(* Logix 5000 project; controller PLC_MCC1300_75F1 vendor 1 type 14 code 166 rev 32.11; software revision 32.04; part 7 of 83 *)

        [109].14   // Speed reference 3 M2CM10S
        [109].15   // Speed reference 4 M2CM10S
        [17].12   // VMCC TD SPARE
        [27].7   // Drive has a fault M2CM01
        [2].3   // VMCC M2 DC Output Power ON
        [113].0   // Drive ready M2CM11S
        [115].0   // Drive ready M2CM11N
        [117].0   // Drive ready M2CM12S
        [119].0   // Drive ready M2CM12N
        [123].11   // MB -->> M2 SPARE
        [31].7   // Drive has a fault M2CM3
        [102]   // RACK 14 INPUT UPDATES
        [104]   // Rack 15 Input Updates
        [1]   // RIO VMCC_TD_Inputs
        [17].13   // VMCC TD SPARE
        [49].11   // PANEL TD-CS4N SPARE
        [123].0   // MB -->> M2 SPARE
        [117].13   // Speed reference 2 M2CM12S
        [17].14   // VMCC TD SPARE
        [3].15   // VMCC M2 Drive fault Reset
        [53].13   // PANEL TD-CS5N SPARE
        [17].8   // VMCC TD Alarm Silence
        [2].10   // VMCC M2 E-STOP ACTIVE
        [2].5   // VMCC M2 E-STOP Power ON
        [32].12   // PANEL KD-CS1N SPARE
        [123].12   // MB -->> M2 SPARE
        [49].12   // PANEL TD-CS4N SPARE
        [106]   // Rack 15 Input Updates
        [108]   // Rack 15 Input Updates
        [17].15   // VMCC TD SPARE
        [49].13   // PANEL TD-CS4N SPARE
        [123].6   // MB -->> M2 SPARE
        [18].10   // VMCC TD SPARE
        [53].14   // PANEL TD-CS5N SPARE
        [53].15   // PANEL TD-CS5N SPARE
        [32].13   // PANEL KD-CS1N SPARE
        [32].14   // PANEL KD-CS1N SPARE
        [32].15   // PANEL KD-CS1N SPARE
        [33].10   // PANEL KD-CS1N SPARE
        [123].13   // MB -->> M2 SPARE
        [49].14   // PANEL TD-CS4N SPARE
        [110]   // Rack 15 Input Updates
        [112]   // Rack 16 Input Updates
        [18].11   // VMCC TD SPARE
        [49].15   // PANEL TD-CS4N SPARE
        [123].7   // MB -->> M2 SPARE
        [1].5   // Rockwell Run out Speed up signal M2CM7
        [117].14   // Speed reference 3 M2CM12S
        [123].8   // MB -->> M2 SPARE
        [117].15   // Speed reference 4 M2CM12S
        [117].2   // Command direction FW M2CM12S
        [117].3   // Actual direction FWD M2CM12S
        [33].0   // PANEL KD-CS1N Trim deck Move IN North Selector Sw.
        [36].2   // PANEL TD-CS1N Trim knocker 1 AUTO South Selector Sw.
        [117].6   // Drive has an alarm M2CM12S
        [117].7   // Drive has a fault M2CM12S
        [18].12   // VMCC TD SPARE
        [56].12   // PANEL TD-CS5S SPARE
        [56].13   // PANEL TD-CS5S SPARE
        [33].11   // PANEL KD-CS1N SPARE
        [33].12   // PANEL KD-CS1N SPARE
        [33].13   // PANEL KD-CS1N SPARE
        [33].14   // PANEL KD-CS1N SPARE
        [123].14   // MB -->> M2 SPARE
        [52].12   // PANEL TD-CS5N SPARE
        [114]   // Rack 16 Input Updates
        [116]   // Rack 16 Input Updates
        [18].13   // VMCC TD SPARE
        [52].13   // PANEL TD-CS5N SPARE
        [123].9   // MB -->> M2 SPARE
        [18].14   // VMCC TD SPARE
        [56].14   // PANEL TD-CS5S SPARE
        [57].10   // PANEL TD-CS5S SPARE
        [33].15   // PANEL KD-CS1N SPARE
        [37].11   // PANEL TD-CS1N SPARE
        [37].12   // PANEL TD-CS1N SPARE
        [37].13   // PANEL TD-CS1N SPARE
        [123].15   // MB -->> M2 SPARE
        [52].14   // PANEL TD-CS5N SPARE
        [118]   // Rack 16 Input Updates
        [120]   // Rack 17 Input Updates
        [18].15   // VMCC TD SPARE
        [52].15   // PANEL TD-CS5N SPARE
        [57].11   // PANEL TD-CS5S SPARE
        [57].12   // PANEL TD-CS5S SPARE
        [37].14   // PANEL TD-CS1N SPARE
        [37].15   // PANEL TD-CS1N SPARE
        [40].12   // PANEL TD-CS2N SPARE
        [40].13   // PANEL TD-CS2N SPARE
        [24].12   // I-SCAN BARS ON/OFF
        [53].10   // PANEL TD-CS5N SPARE
        [17].9   // VMCC TD Alarm Reset
        [29].1   // Drive running M2CM2
        [53].11   // PANEL TD-CS5N SPARE
        [1].6   // Rockwell Run out Speed up signal M2CM8
        [73].5   // BENCHBOARD Knurl Knocker Nth & Sth Auto mode
        [64].12   // Trim Deck PANEL TD-CS3S Crush all OFF Switch
        [73].7   // BENCHBOARD Knurl Knocker Master Auto mode
        [1].7   // Rockwell Run out Speed up signal M2CM9
        [37].7   // PANEL TD-CS1N Trim Conv 1 North Outer Limit Sw.
        [37].8   // PANEL TD-CS1N Trim Conv 1 North Inner Limit Sw.
        [33].8   // PANEL KD-CS1N Trim deck South Outer Limit Sw.
        [24].3   // RELIANCE CAPPING SYSTEM Trim Knocker #2 North Lower wheel
        [72].6   // BENCHBOARD Trim knocker #2 South Up Selector Sw.
        [72].8   // BENCHBOARD Trim knocker #3 North Up Selector Sw.
        [73].0   // BENCHBOARD Trim knocker #5 North Up Selector Sw.
        [24].15   // RELIANCE CAPPING SYSTEM Tracking window Lamp ON
        [33].4   // PANEL KD-CS1N Knurl knocker North Outer Limit Sw.
        [33].5   // PANEL KD-CS1N Knurl knocker North Inner Limit Sw.
        [33].9   // PANEL KD-CS1N Trim deck South Inner Limit Sw.
        [24].4   // RELIANCE CAPPING SYSTEM Trim Knocker #2 South Lower wheel
        [73].2   // BENCHBOARD Trim knocker #5 South Up Selector Sw.
        [37].10   // PANEL TD-CS1N Trim Conv 1 South Inner Limit Sw.
        [41].10   // PANEL TD-CS2N Trim Conv 2 North Outer Limit Sw.
        [41].11   // PANEL TD-CS2N Trim Conv 2 North Inner Limit Sw.
        [4].11   // VMCC M2 Speed zone 12 Drive Fault * 2CM12N
        [72].1   // BENCHBOARD Trim knocker #5 North Auto mode
        [72].3   // BENCHBOARD Trim knocker #5 South Auto mode
        [36].12   // PANEL TD-CS1N Float Glass Hold Down Wheels Auto Sel. Sw.
        [24].0   // RELIANCE CAPPING SYSTEM Knurl Knocker Nth & Sth Lower wheel
        [32].4   // PANEL KD-CS1N Knurl knocker Move UP South Selector Sw.
        [125].2   // ROCKWELL CAPPER Input to Disable manual y-cut bar 1
        [37].9   // PANEL TD-CS1N Trim Conv 1 South Outer Limit Sw.
        [36].1   // PANEL TD-CS1N Trim knocker 1 Move OUT South Selector Sw.
        [36].4   // PANEL TD-CS1N Trim knocker 1 Move UP South Selector Sw.
        [24].10   // RELIANCE CAPPING SYSTEM Trim Knocker #5 South Lower wheel
        [44].13   // Trim Deck PANEL TD-CS3N Crush all ON Switch
        [72].7   // BENCHBOARD Trim knocker #2 South Auto mode
        [45].6   // PANEL TD-CS3N Trim Conv 3 North Outer Limit Sw.
        [32].6   // PANEL KD-CS1N Knurl knocker Move IN North Selector Sw.
        [45].7   // PANEL TD-CS3N Trim Conv 3 North Inner Limit Sw.
        [72].9   // BENCHBOARD Trim knocker #3 North Auto mode
        [40].10   // PANEL TD-CS2N Trim knocker #2 Move UP North Selector Sw.
        [24].5   // RELIANCE CAPPING SYSTEM Trim Knocker #3 North Lower wheel
        [88]   // RACK 13 INPUT UPDATES
        [74]   // RACK 7 INPUT UPDATES
        [40].14   // PANEL TD-CS2N SPARE
        [24].6   // RELIANCE CAPPING SYSTEM Trim Knocker #3 South Lower wheel
        [90]   // RACK 13 INPUT UPDATES
        [103].14   // Speed reference 3 M2CM8N
        [119].10   // Local control 2 M2CM12N
        [109].2   // Command direction FW M2CM10S
        [115].12   // Speed reference 1 M2CM11N
        [36].8   // PANEL TD-CS1N Trim knocker 1 AUTO North Selector Sw.
        [36].14   // PANEL TD-CS1N Eclipse Hold Down Wheels Auto Sel. Sw.
        [36].3   // PANEL TD-CS1N Trim knocker 1 MANUAL South Selector Sw.
        [36].9   // PANEL TD-CS1N Trim knocker 1 MANUAL North Selector Sw.
        [69].5   // PANEL TD-CS2S Trim Conv 2 Move OUT North Selector Sw.
        [125].3   // ROCKWELL CAPPER Input to Disable auto y-cut bar 4
        [56].6   // PANEL TD-CS5S Trim knocker #5 Move IN North Selector Sw.
        [18].3   // VMCC TD SPARE
        [40].15   // PANEL TD-CS2N SPARE
        [41].14   // PANEL TD-CS2N SPARE
        [107].11   // Local control 3 M2CM9N
        [107].6   // Drive has an alarm M2CM9N
        [107].7   // Drive has a fault M2CM9N
        [105].9   // Local control 1 M2CM9S
        [41].15   // PANEL TD-CS2N SPARE
        [109].4   // Accelerating M2CM10S
        [2].8   // VMCC M2 Alarm Silence
        [31].1   // Drive running M2CM3
        [27].1   // Drive running M2CM01
        [18].5   // VMCC TD SPARE
        [44].14   // PANEL TD-CS3N SPARE
        [44].15   // PANEL TD-CS3N SPARE
        [109].10   // Local control 2 M2CM10S
        [109].11   // Local control 3 M2CM10S
        [109].7   // Drive has a fault M2CM10S
        [107].9   // Local control 1 M2CM9N
        [45].10   // PANEL TD-CS3N SPARE
        [109].5   // Decelerating M2CM10S
        [37].0   // PANEL TD-CS1N SPARE
        [37].1   // PANEL TD-CS1N SPARE
        [85].1   // Drive running M2CM4S
        [109].8   // Drive at speed M2CM10S
        [18].6   // VMCC TD SPARE
        [45].11   // PANEL TD-CS3N SPARE
        [45].12   // PANEL TD-CS3N SPARE
        [111].10   // Local control 2 M2CM10N
        [111].11   // Local control 3 M2CM10N
        [111].7   // Drive has a fault M2CM10N
        [111].8   // Drive at speed M2CM10N
        [45].13   // PANEL TD-CS3N SPARE
        [111].4   // Accelerating M2CM10N
        [37].4   // PANEL TD-CS1N SPARE
        [37].5   // PANEL TD-CS1N SPARE
        [87].1   // Drive running M2CM4N
        [18].7   // VMCC TD SPARE
        [45].14   // PANEL TD-CS3N SPARE
        [45].15   // PANEL TD-CS3N SPARE
        [113].10   // Local control 2 M2CM11S
        [113].11   // Local control 3 M2CM11S
        [113].7   // Drive has a fault M2CM11S
        [113].8   // Drive at speed M2CM11S
        [48].12   // PANEL TD-CS4N SPARE
        [111].5   // Decelerating M2CM10N
        [37].6   // PANEL TD-CS1N SPARE
        [4].12   // VMCC M2 Drive alarm
        [89].1   // Drive running M2CM5S
        [33].2   // PANEL KD-CS1N Trim deck Move IN South Selector Sw.
        [32].3   // PANEL KD-CS1N Knurl knocker MANUAL South Selector Sw.
        [73].14   // BENCHBOARD Input Power ON
        [57].13   // PANEL TD-CS5S SPARE
        [41].12   // PANEL TD-CS2N Trim Conv 2 South Outer Limit Sw.
        [36].11   // PANEL TD-CS1N Trim knocker 1 Move DOWN North Selector Sw.
        [3].9   // VMCC M2 Speed zone 10 Drive Fault 2CM10S
        [4].0   // VMCC M2 Speed zone 1 Drive Fault * 2CM01
        [4].1   // VMCC M2 Speed zone 2 Drive Fault * 2CM02
        [4].2   // VMCC M2 Speed zone 3 Drive Fault * 2CM03
        [73].3   // BENCHBOARD Knocker #5 South Auto mode
        [3].6   // VMCC M2 Speed zone 7 Drive Fault * 2CM07S
        [73].10   // Reliance BENCHBOARD Crush all OFF Switch
        [53].12   // PANEL TD-CS5N SPARE
        [113].4   // Accelerating M2CM11S
        [115].8   // Drive at speed M2CM11N
        [48].13   // PANEL TD-CS4N SPARE
        [73].15   // BENCHBOARD Output Power ON
        [117].8   // Drive at speed M2CM12S
        [36].13   // PANEL TD-CS1N Float Glass Hold Down Wheels Up Sel. Sw.
        [68].0   // PANEL TD-CS2S Trim knocker #2 Move IN South Selector Sw.
        [115].13   // Speed reference 2 M2CM11N
        [76].12   // PANEL KD-CS1S SPARE
        [40].5   // PANEL TD-CS2N Trim knocker #2 Move DOWN South Selector Sw.
        [44].10   // PANEL TD-CS3N Trim knocker #3 Move UP North Selector Sw.
        [44].5   // PANEL TD-CS3N Trim knocker #3 Move DOWN South Selector Sw.
        [24].7   // RELIANCE CAPPING SYSTEM Trim Knocker #4 North Lower wheel
        [103].2   // Command direction FW M2CM8N
        [125].4   // ROCKWELL CAPPER Input to Disable auto y-cut bar 3
        [103].15   // Speed reference 4 M2CM8N
        [2].0   // VMCC TD SPARE
        [81].0   // PANEL TD-CS1S SPARE
        [81].1   // PANEL TD-CS1S SPARE
        [57].14   // PANEL TD-CS5S SPARE
        [57].15   // PANEL TD-CS5S SPARE
        [60].12   // PANEL TD-CS4S SPARE
        [113].5   // Decelerating M2CM11S
        [81].4   // PANEL TD-CS1S SPARE
        [91].1   // Drive running M2CM5N
        [92]   // RACK 13 INPUT UPDATES
        [94]   // RACK 13 INPUT UPDATES
        [18].8   // VMCC TD SPARE
        [18].9   // VMCC TD SPARE
        [2].4   // VMCC M2 SPARE
        [81].5   // PANEL TD-CS1S SPARE
        [81].6   // PANEL TD-CS1S SPARE
        [60].13   // PANEL TD-CS4S SPARE
        [60].14   // PANEL TD-CS4S SPARE
        [60].15   // PANEL TD-CS4S SPARE
        [115].4   // Accelerating M2CM11N
        [93].1   // Drive running M2CM6S
        [96]   // RACK 14 INPUT UPDATES
        [98]   // RACK 14 INPUT UPDATES
        [2].13   // VMCC M2 SPARE
        [2].14   // VMCC M2 SPARE
        [3].0   // VMCC M2 SPARE
        [61].10   // PANEL TD-CS4S SPARE
        [61].11   // PANEL TD-CS4S SPARE
        [61].12   // PANEL TD-CS4S SPARE
        [115].5   // Decelerating M2CM11N
        [95].1   // Drive running M2CM6N
        [2].15   // VMCC M2 SPARE
        [3].12   // VMCC M2 SPARE
        [3].1   // VMCC M2 SPARE
        [61].13   // PANEL TD-CS4S SPARE
        [61].14   // PANEL TD-CS4S SPARE
        [61].15   // PANEL TD-CS4S SPARE
        [117].4   // Accelerating M2CM12S
        [97].1   // Drive running M2CM7S
        [3].13   // VMCC M2 SPARE
        [3].14   // VMCC M2 SPARE
        [3].2   // VMCC M2 SPARE
        [64].14   // PANEL TD-CS3S SPARE
        [64].15   // PANEL TD-CS3S SPARE
        [65].10   // PANEL TD-CS3S SPARE
        [117].5   // Decelerating M2CM12S
        [99].1   // Drive running M2CM7N
        [4].13   // VMCC M2 SPARE
        [4].14   // VMCC M2 SPARE
        [3].7   // VMCC M2 Speed zone 8 Drive Fault * 2CM08S
        [65].11   // PANEL TD-CS3S SPARE
        [65].12   // PANEL TD-CS3S SPARE
        [65].13   // PANEL TD-CS3S SPARE
        [119].4   // Accelerating M2CM12N
        [4].15   // VMCC M2 SPARE
        [64].13   // Trim Deck PANEL TD-CS3S Crush all ON Switch
        [41].13   // PANEL TD-CS2N Trim Conv 2 South Inner Limit Sw.
        [77].6   // PANEL KD-CS1S Trim deck North Outer Limit Sw.
        [45].8   // PANEL TD-CS3N Trim Conv 3 South Outer Limit Sw.
        [36].7   // PANEL TD-CS1N Trim knocker 1 Move OUT North Selector Sw.
        [69].10   // PANEL TD-CS2S Trim Conv 2 North Outer Limit Sw.
        [41].0   // PANEL TD-CS2N Trim Conv 1 Move IN North Selector Sw.
        [48].10   // PANEL TD-CS4N Trim knocker #4 Move UP North Selector Sw.
        [109].3   // Actual direction FWD M2CM10S
        [76].13   // PANEL KD-CS1S SPARE
        [109].6   // Drive has an alarm M2CM10S
        [40].0   // PANEL TD-CS2N Trim knocker #2 Move IN South Selector Sw.
        [32].9   // PANEL KD-CS1N Knurl knocker MANUAL North Selector Sw.
        [40].4   // PANEL TD-CS2N Trim knocker #2 Move UP South Selector Sw.
        [68].1   // PANEL TD-CS2S Trim knocker #2 Move OUT South Selector Sw.
        [52].1   // PANEL TD-CS5N Trim knocker #5 Move OUT South Selector Sw.
        [115].14   // Speed reference 3 M2CM11N
        [24].8   // RELIANCE CAPPING SYSTEM Trim Knocker #4 South Lower wheel
        [45].9   // PANEL TD-CS3N Trim Conv 3 South Inner Limit Sw.
        [69].7   // PANEL TD-CS2S Trim Conv 2 Move OUT South Selector Sw.
        [52].10   // PANEL TD-CS5N Trim knocker #5 Move UP North Selector Sw.
        [24].9   // RELIANCE CAPPING SYSTEM Trim Knocker #5 North Lower wheel
        [119].11   // Local control 3 M2CM12N
        [65].14   // PANEL TD-CS3S SPARE
        [76].14   // PANEL KD-CS1S SPARE
        [103].3   // Actual direction FWD M2CM8N
        [105].13   // Speed reference 2 M2CM9S
        [105].14   // Speed reference 3 M2CM9S
        [111].12   // Speed reference 1 M2CM10N
        [76].7   // PANEL KD-CS1S Knurl knocker Move OUT North Selector Sw.
        [80].0   // PANEL TD-CS1S Trim knocker 1 Move IN South Selector Sw.
        [119].12   // Speed reference 1 M2CM12N
        [105].15   // Speed reference 4 M2CM9S
        [111].13   // Speed reference 2 M2CM10N
        [119].13   // Speed reference 2 M2CM12N
        [40].11   // PANEL TD-CS2N Trim knocker #2 Move DOWN North Selector Sw.
        [56].7   // PANEL TD-CS5S Trim knocker #5 Move OUT North Selector Sw.
        [44].11   // PANEL TD-CS3N Trim knocker #3 Move DOWN North Selector Sw.
        [60].0   // PANEL TD-CS4S Trim knocker #4 Move IN South Selector Sw.
        [36].10   // PANEL TD-CS1N Trim knocker 1 Move UP North Selector Sw.
        [48].11   // PANEL TD-CS4N Trim knocker #4 Move DOWN North Selector Sw.
        [48].14   // PANEL TD-CS4N SPARE
        [105].12   // Speed reference 1 M2CM9S
        [69].11   // PANEL TD-CS2S Trim Conv 2 North Inner Limit Sw.
        [49].6   // PANEL TD-CS4N Trim Conv 4 North Outer Limit Sw.
        [48].15   // PANEL TD-CS4N SPARE
        [49].10   // PANEL TD-CS4N SPARE
        [60].1   // PANEL TD-CS4S Trim knocker #4 Move OUT South Selector Sw.
        [60].10   // PANEL TD-CS4S Trim knocker #4 Move UP North Selector Sw.
        [60].11   // PANEL TD-CS4S Trim knocker #4 Move DOWN North Selector Sw.
        [60].4   // PANEL TD-CS4S Trim knocker #4 Move UP South Selector Sw.
        [60].5   // PANEL TD-CS4S Trim knocker #4 Move DOWN South Selector Sw.
        [60].6   // PANEL TD-CS4S Trim knocker #4 Move IN North Selector Sw.
        [60].7   // PANEL TD-CS4S Trim knocker #4 Move OUT North Selector Sw.
        [76].15   // PANEL KD-CS1S SPARE
        [77].10   // PANEL KD-CS1S SPARE
        [77].11   // PANEL KD-CS1S SPARE
        [77].12   // PANEL KD-CS1S SPARE
        [77].13   // PANEL KD-CS1S SPARE
        [77].14   // PANEL KD-CS1S SPARE
        [77].15   // PANEL KD-CS1S SPARE
        [81].11   // PANEL TD-CS1S SPARE
        [81].12   // PANEL TD-CS1S SPARE
        [81].13   // PANEL TD-CS1S SPARE
        [81].14   // PANEL TD-CS1S SPARE
        [52].4   // PANEL TD-CS5N Trim knocker #5 Move UP South Selector Sw.
        [48].4   // PANEL TD-CS4N Trim knocker #4 Move UP South Selector Sw.
        [48].5   // PANEL TD-CS4N Trim knocker #4 Move DOWN South Selector Sw.
        [48].6   // PANEL TD-CS4N Trim knocker #4 Move IN North Selector Sw.
        [80].1   // PANEL TD-CS1S Trim knocker 1 Move OUT South Selector Sw.
        [41].2   // PANEL TD-CS2N Trim Conv 1 Move IN South Selector Sw.
        [40].2   // PANEL TD-CS2N Trim knocker #2 AUTO South Selector Sw.
        [40].8   // PANEL TD-CS2N Trim knocker #2 AUTO North Selector Sw.
        [119].14   // Speed reference 3 M2CM12N
        [69].12   // PANEL TD-CS2S Trim Conv 2 South Outer Limit Sw.
        [3].8   // VMCC M2 Speed zone 9 Drive Fault * 2CM09S
        [69].13   // PANEL TD-CS2S Trim Conv 2 South Inner Limit Sw.
        [4].3   // VMCC M2 Speed zone 4 Drive Fault * 2CM04N
        [77].4   // PANEL KD-CS1S Knurl knocker South Outer Limit Sw.
        [77].5   // PANEL KD-CS1S Knurl knocker South Inner Limit Sw.
        [4].4   // VMCC M2 Speed zone 5 Drive Fault * 2CM05N
        [80].15   // PANEL TD-CS1S Eclipse Hold Down Wheels Sel. Sw.
        [81].10   // PANEL TD-CS1S Trim Conv 1 South Inner Limit Sw.
        [4].5   // VMCC M2 Speed zone 6 Drive Fault * 2CM06N
        [4].6   // VMCC M2 Speed zone 7 Drive Fault * 2CM07N
        [4].7   // VMCC M2 Speed zone 8 Drive Fault * 2CM08N
        [4].8   // VMCC M2 Speed zone 9 Drive Fault * 2CM09N
        [4].9   // VMCC M2 Speed zone 10 Drive Fault * 2CM10
        [41].4   // PANEL TD-CS2N Trim Conv 2 Move IN North Selector Sw.
        [36].6   // PANEL TD-CS1N Trim knocker 1 Move IN North Selector Sw.
        [41].6   // PANEL TD-CS2N Trim Conv 2 Move IN South Selector Sw.
        [80].4   // PANEL TD-CS1S Trim knocker 1 Move UP South Selector Sw.
        [45].0   // PANEL TD-CS3N Trim Conv 3 Move IN North Selector Sw.
        [37].2   // PANEL TD-CS1N Trim knocker 1 North Outer Limit Sw.
        [40].3   // PANEL TD-CS2N Trim knocker #2 MANUAL South Selector Sw.
        [80].5   // PANEL TD-CS1S Trim knocker 1 Move DOWN South Selector Sw.
        [45].2   // PANEL TD-CS3N Trim Conv 3 Move IN South Selector Sw.
        [37].3   // PANEL TD-CS1N Trim knocker 1 North Inner Limit Sw.
        [49].0   // PANEL TD-CS4N Trim Conv 4 Move IN North Selector Sw.
        [72].10   // BENCHBOARD Trim knocker #3 South Up Selector Sw.
        [49].2   // PANEL TD-CS4N Trim Conv 4 Move IN South Selector Sw.
        [72].12   // BENCHBOARD Trim knocker #4 North Up Selector Sw.
        [53].0   // PANEL TD-CS5N Trim Conv 5 Move IN North Selector Sw.
        [72].14   // BENCHBOARD Trim knocker #4 South Up Selector Sw.
        [53].2   // PANEL TD-CS5N Trim Conv 5 Move IN South Selector Sw.
        [73].4   // BENCHBOARD Knurl Knocker Nth & Sth Up Selector Sw.
        [57].0   // PANEL TD-CS5S Trim Conv 5 Move IN North Selector Sw.
        [52].5   // PANEL TD-CS5N Trim knocker #5 Move DOWN South Selector Sw.
        [77].0   // PANEL KD-CS1S Trim deck Move IN North Selector Sw.
        [48].7   // PANEL TD-CS4N Trim knocker #4 Move OUT North Selector Sw.
        [40].9   // PANEL TD-CS2N Trim knocker #2 MANUAL North Selector Sw.
        [68].10   // PANEL TD-CS2S Trim knocker #2 Move UP North Selector Sw.
        [77].2   // PANEL KD-CS1S Trim deck Move IN South Selector Sw.
        [80].10   // PANEL TD-CS1S Trim knocker 1 Move UP North Selector Sw.
        [81].2   // PANEL TD-CS1S Trim knocker 1 South Outer Limit Sw.
        [57].2   // PANEL TD-CS5S Trim Conv 5 Move IN South Selector Sw.
        [52].11   // PANEL TD-CS5N Trim knocker #5 Move DOWN North Selector Sw.
        [56].1   // PANEL TD-CS5S Trim knocker #5 Move OUT South Selector Sw.
        [64].0   // PANEL TD-CS3S Trim knocker #3 Move IN South Selector Sw.
        [64].1   // PANEL TD-CS3S Trim knocker #3 Move OUT South Selector Sw.
        [64].10   // PANEL TD-CS3S Trim knocker #3 Move UP North Selector Sw.
        [64].11   // PANEL TD-CS3S Trim knocker #3 Move DOWN North Selector Sw.
        [36].5   // PANEL TD-CS1N Trim knocker 1 Move DOWN South Selector Sw.
        [119].15   // Speed reference 4 M2CM12N
        [40].1   // PANEL TD-CS2N Trim knocker #2 Move OUT South Selector Sw.
        [41].1   // PANEL TD-CS2N Trim Conv 1 Move OUT North Selector Sw.
        [41].3   // PANEL TD-CS2N Trim Conv 1 Move OUT South Selector Sw.
        [41].5   // PANEL TD-CS2N Trim Conv 2 Move OUT North Selector Sw.
        [41].7   // PANEL TD-CS2N Trim Conv 2 Move OUT South Selector Sw.
        [44].2   // PANEL TD-CS3N Trim knocker #3 AUTO South Selector Sw.
        [44].8   // PANEL TD-CS3N Trim knocker #3 AUTO North Selector Sw.
        [45].1   // PANEL TD-CS3N Trim Conv 3 Move OUT North Selector Sw.
        [52].6   // PANEL TD-CS5N Trim knocker #5 Move IN North Selector Sw.
        [64].4   // PANEL TD-CS3S Trim knocker #3 Move UP South Selector Sw.
        [64].5   // PANEL TD-CS3S Trim knocker #3 Move DOWN South Selector Sw.
        [40].7   // PANEL TD-CS2N Trim knocker #2 Move OUT North Selector Sw.
        [64].6   // PANEL TD-CS3S Trim knocker #3 Move IN North Selector Sw.
        [52].7   // PANEL TD-CS5N Trim knocker #5 Move OUT North Selector Sw.
        [44].3   // PANEL TD-CS3N Trim knocker #3 MANUAL South Selector Sw.
        [61].0   // PANEL TD-CS4S Trim Conv 4 Move IN North Selector Sw.
        [80].11   // PANEL TD-CS1S Trim knocker 1 Move DOWN North Selector Sw.
        [56].10   // PANEL TD-CS5S Trim knocker #5 Move UP North Selector Sw.
        [80].6   // PANEL TD-CS1S Trim knocker 1 Move IN North Selector Sw.
        [68].11   // PANEL TD-CS2S Trim knocker #2 Move DOWN North Selector Sw.
        [56].0   // PANEL TD-CS5S Trim knocker #5 Move IN South Selector Sw.
        [44].9   // PANEL TD-CS3N Trim knocker #3 MANUAL North Selector Sw.
        [81].15   // PANEL TD-CS1S SPARE
        [61].2   // PANEL TD-CS4S Trim Conv 4 Move IN South Selector Sw.
        [65].0   // PANEL TD-CS3S Trim Conv 3 Move IN North Selector Sw.
        [64].7   // PANEL TD-CS3S Trim knocker #3 Move OUT North Selector Sw.
        [56].11   // PANEL TD-CS5S Trim knocker #5 Move DOWN North Selector Sw.
        [80].12   // PANEL TD-CS1S Float Glass Hold Down Wheels Auto Sel. Sw.
        [45].3   // PANEL TD-CS3N Trim Conv 3 Move OUT South Selector Sw.
        [80].13   // PANEL TD-CS1S Float Glass Hold Down Wheels Up Sel. Sw.
        [68].4   // PANEL TD-CS2S Trim knocker #2 Move UP South Selector Sw.
        [80].7   // PANEL TD-CS1S Trim knocker 1 Move OUT North Selector Sw.
        [49].7   // PANEL TD-CS4N Trim Conv 4 North Inner Limit Sw.
        [49].8   // PANEL TD-CS4N Trim Conv 4 South Outer Limit Sw.
        [49].9   // PANEL TD-CS4N Trim Conv 4 South Inner Limit Sw.
        [53].6   // PANEL TD-CS5N Trim Conv 5 North Outer Limit Sw.
        [53].7   // PANEL TD-CS5N Trim Conv 5 North Inner Limit Sw.
        [57].6   // PANEL TD-CS5S Trim Conv 5 North Outer Limit Sw.
        [57].7   // PANEL TD-CS5S Trim Conv 5 North Inner Limit Sw.
        [57].8   // PANEL TD-CS5S Trim Conv 5 South Outer Limit Sw.
        [57].9   // PANEL TD-CS5S Trim Conv 5 South Inner Limit Sw.
        [61].6   // PANEL TD-CS4S Trim Conv 4 North Outer Limit Sw.
        [81].3   // PANEL TD-CS1S Trim knocker 1 South Inner Limit Sw.
        [119].2   // Command direction FW M2CM12N
        [85].7   // Drive has a fault M2CM4S
        [44].1   // PANEL TD-CS3N Trim knocker #3 Move OUT South Selector Sw.
        [61].7   // PANEL TD-CS4S Trim Conv 4 North Inner Limit Sw.
        [61].8   // PANEL TD-CS4S Trim Conv 4 South Outer Limit Sw.
        [48].3   // PANEL TD-CS4N Trim knocker #4 MANUAL South Selector Sw.
        [48].2   // PANEL TD-CS4N Trim knocker #4 AUTO South Selector Sw.
        [87].7   // Drive has a fault M2CM4N
        [61].9   // PANEL TD-CS4S Trim Conv 4 South Inner Limit Sw.
        [89].7   // Drive has a fault M2CM5S
        [68].5   // PANEL TD-CS2S Trim knocker #2 Move DOWN South Selector Sw.
        [48].8   // PANEL TD-CS4N Trim knocker #4 AUTO North Selector Sw.
        [65].6   // PANEL TD-CS3S Trim Conv 3 North Outer Limit Sw.
        [119].3   // Actual direction FWD M2CM12N
        [68].6   // PANEL TD-CS2S Trim knocker #2 Move IN North Selector Sw.
        [65].2   // PANEL TD-CS3S Trim Conv 3 Move IN South Selector Sw.
        [44].6   // PANEL TD-CS3N Trim knocker #3 Move IN North Selector Sw.
        [40].6   // PANEL TD-CS2N Trim knocker #2 Move IN North Selector Sw.
        [119].6   // Drive has an alarm M2CM12N
        [44].0   // PANEL TD-CS3N Trim knocker #3 Move IN South Selector Sw.
        [68].7   // PANEL TD-CS2S Trim knocker #2 Move OUT North Selector Sw.
        [69].0   // PANEL TD-CS2S Trim Conv 1 Move IN North Selector Sw.
        [44].7   // PANEL TD-CS3N Trim knocker #3 Move OUT North Selector Sw.
        [65].7   // PANEL TD-CS3S Trim Conv 3 North Inner Limit Sw.
        [65].8   // PANEL TD-CS3S Trim Conv 3 South Outer Limit Sw.
        [65].9   // PANEL TD-CS3S Trim Conv 3 South Inner Limit Sw.
        [73].6   // BENCHBOARD Knurl Knocker Master Up Selector Sw.
        [81].7   // PANEL TD-CS1S Trim Conv 1 North Outer Limit Sw.
        [81].8   // PANEL TD-CS1S Trim Conv 1 North Inner Limit Sw.
        [81].9   // PANEL TD-CS1S Trim Conv 1 South Outer Limit Sw.
        [48].0   // PANEL TD-CS4N Trim knocker #4 Move IN South Selector Sw.
        [77].7   // PANEL KD-CS1S Trim deck North Inner Limit Sw.
        [77].8   // PANEL KD-CS1S Trim deck South Outer Limit Sw.
        [77].9   // PANEL KD-CS1S Trim deck South Inner Limit Sw.
        [52].0   // PANEL TD-CS5N Trim knocker #5 Move IN South Selector Sw.
        [91].7   // Drive has a fault M2CM5N
        [93].7   // Drive has a fault M2CM6S
        [95].7   // Drive has a fault M2CM6N
        [97].7   // Drive has a fault M2CM7S
        [69].2   // PANEL TD-CS2S Trim Conv 1 Move IN South Selector Sw.
        [56].4   // PANEL TD-CS5S Trim knocker #5 Move UP South Selector Sw.
        [49].1   // PANEL TD-CS4N Trim Conv 4 Move OUT North Selector Sw.
        [125].5   // ROCKWELL CAPPER Input to Disable auto y-cut bar 2
        [125].6   // ROCKWELL CAPPER Input to Disable auto y-cut bar 1
        [32].2   // PANEL KD-CS1N Knurl knocker AUTO South Selector Sw.
        [32].8   // PANEL KD-CS1N Knurl knocker AUTO North Selector Sw.
        [33].1   // PANEL KD-CS1N Trim deck Move OUT North Selector Sw.
        [33].3   // PANEL KD-CS1N Trim deck Move OUT South Selector Sw.
        [41].8   // PANEL TD-CS2N Trim knocker #2 North Outer Limit Sw.
        [41].9   // PANEL TD-CS2N Trim knocker #2 North Inner Limit Sw.
        [45].4   // PANEL TD-CS3N Trim knocker #3 North Outer Limit Sw.
        [45].5   // PANEL TD-CS3N Trim knocker #3 North Inner Limit Sw.
        [49].4   // PANEL TD-CS4N Trim knocker #4 North Outer Limit Sw.
        [49].5   // PANEL TD-CS4N Trim knocker #4 North Inner Limit Sw.
        [53].8   // PANEL TD-CS5S Trim knocker #5 South Outer Limit Sw.
        [53].9   // PANEL TD-CS5S Trim knocker #5 South Inner Limit Sw.
        [61].4   // PANEL TD-CS4S Trim knocker #4 South Outer Limit Sw.
        [61].5   // PANEL TD-CS4S Trim knocker #4 South Inner Limit Sw.
        [65].4   // PANEL TD-CS3S Trim knocker #3 South Outer Limit Sw.
        [99].7   // Drive has a fault M2CM7N
        [119].7   // Drive has a fault M2CM12N
        [17].11   // VMCC TD Panel Overtemp Alarm
        [17].3   // VMCC TD DC Output Power ON
        [17].4   // VMCC TD DC Power Supply #1 ON
        [76].10   // PANEL KD-CS1S Knurl knocker Move UP North Selector Sw.
        [49].3   // PANEL TD-CS4N Trim Conv 4 Move OUT South Selector Sw.
        [76].0   // PANEL KD-CS1S Knurl knocker Move IN South Selector Sw.
        [76].3   // PANEL KD-CS1S Knurl knocker MANUAL South Selector Sw.
        [76].4   // PANEL KD-CS1S Knurl knocker Move UP South Selector Sw.
        [76].6   // PANEL KD-CS1S Knurl knocker Move IN North Selector Sw.
        [17].6   // VMCC TD DC Power Supply #2 ON
        [52].2   // PANEL TD-CS5N Trim knocker #5 AUTO South Selector Sw.
        [52].8   // PANEL TD-CS5N Trim knocker #5 AUTO North Selector Sw.
        [69].4   // PANEL TD-CS2S Trim Conv 2 Move IN North Selector Sw.
        [65].5   // PANEL TD-CS3S Trim knocker #3 South Inner Limit Sw.
        [69].8   // PANEL TD-CS2S Trim knocker #2 South Outer Limit Sw.
        [53].1   // PANEL TD-CS5N Trim Conv 5 Move OUT North Selector Sw.
        [53].3   // PANEL TD-CS5N Trim Conv 5 Move OUT South Selector Sw.
        [69].6   // PANEL TD-CS2S Trim Conv 2 Move IN South Selector Sw.
        [69].9   // PANEL TD-CS2S Trim knocker #2 South Inner Limit Sw.
        [76].2   // PANEL KD-CS1S Knurl knocker AUTO South Selector Sw.
        [56].2   // PANEL TD-CS5S Trim knocker #5 AUTO South Selector Sw.
        [56].8   // PANEL TD-CS5S Trim knocker #5 AUTO North Selector Sw.
        [80].2   // PANEL TD-CS1S Trim knocker 1 AUTO South Selector Sw.
        [76].8   // PANEL KD-CS1S Knurl knocker AUTO North Selector Sw.
        [77].1   // PANEL KD-CS1S Trim deck Move OUT North Selector Sw.
        [57].1   // PANEL TD-CS5S Trim Conv 5 Move OUT North Selector Sw.
        [57].3   // PANEL TD-CS5S Trim Conv 5 Move OUT South Selector Sw.
        [80].8   // PANEL TD-CS1S Trim knocker 1 AUTO North Selector Sw.
        [77].3   // PANEL KD-CS1S Trim deck Move OUT South Selector Sw.
        [48].9   // PANEL TD-CS4N Trim knocker #4 MANUAL North Selector Sw.
        [52].3   // PANEL TD-CS5N Trim knocker #5 MANUAL South Selector Sw.
        [76].9   // PANEL KD-CS1S Knurl knocker MANUAL North Selector Sw.
        [60].2   // PANEL TD-CS4S Trim knocker #4 AUTO South Selector Sw.
        [60].8   // PANEL TD-CS4S Trim knocker #4 AUTO North Selector Sw.
        [52].9   // PANEL TD-CS5N Trim knocker #5 MANUAL North Selector Sw.
        [56].3   // PANEL TD-CS5S Trim knocker #5 MANUAL South Selector Sw.
        [80].14   // PANEL TD-CS1S Eclipse Hold Down Wheels Auto Sel. Sw.
        [61].1   // PANEL TD-CS4S Trim Conv 4 Move OUT North Selector Sw.
        [61].3   // PANEL TD-CS4S Trim Conv 4 Move OUT South Selector Sw.
        [56].9   // PANEL TD-CS5S Trim knocker #5 MANUAL North Selector Sw.
        [60].3   // PANEL TD-CS4S Trim knocker #4 MANUAL South Selector Sw.
        [80].3   // PANEL TD-CS1S Trim knocker 1 MANUAL South Selector Sw.
        [64].2   // PANEL TD-CS3S Trim knocker #3 AUTO South Selector Sw.
        [64].8   // PANEL TD-CS3S Trim knocker #3 AUTO North Selector Sw.
        [60].9   // PANEL TD-CS4S Trim knocker #4 MANUAL North Selector Sw.
        [64].3   // PANEL TD-CS3S Trim knocker #3 MANUAL South Selector Sw.
        [80].9   // PANEL TD-CS1S Trim knocker 1 MANUAL North Selector Sw.
        [65].1   // PANEL TD-CS3S Trim Conv 3 Move OUT North Selector Sw.
        [65].3   // PANEL TD-CS3S Trim Conv 3 Move OUT South Selector Sw.
        [64].9   // PANEL TD-CS3S Trim knocker #3 MANUAL North Selector Sw.
        [68].3   // PANEL TD-CS2S Trim knocker #2 MANUAL South Selector Sw.
        [68].2   // PANEL TD-CS2S Trim knocker #2 AUTO South Selector Sw.
        [68].8   // PANEL TD-CS2S Trim knocker #2 AUTO North Selector Sw.
        [68].9   // PANEL TD-CS2S Trim knocker #2 MANUAL North Selector Sw.
        [76].1   // PANEL KD-CS1S Knurl knocker Move OUT South Selector Sw.
        [69].1   // PANEL TD-CS2S Trim Conv 1 Move OUT North Selector Sw.
        [69].3   // PANEL TD-CS2S Trim Conv 1 Move OUT South Selector Sw.
        [44].4   // PANEL TD-CS3N Trim knocker #3 Move UP South Selector Sw.
        [17].7   // VMCC TD DC Power Supply #3 ON
        [48].1   // PANEL TD-CS4N Trim knocker #4 Move OUT South Selector Sw.
   KD_N_MOVIN : ALIAS FOR N14[256].0;
   KD_N_MOVOUT : ALIAS FOR N14[257].0;
   KD_S_MOVIN : ALIAS FOR N14[256].1;
   KD_S_MOVOUT : ALIAS FOR N14[257].1;
   KK_N_MOVDN : ALIAS FOR N14[253].0;
   KK_N_MOVIN : ALIAS FOR N14[254].0;
   KK_N_MOVOUT : ALIAS FOR N14[255].0;
   KK_N_MOVUP : ALIAS FOR N14[252].0;
   KK_S_MOVDN : ALIAS FOR N14[253].1;
   KK_S_MOVIN : ALIAS FOR N14[254].1;
   KK_S_MOVOUT : ALIAS FOR N14[255].1;
   KK_S_MOVUP : ALIAS FOR N14[252].1;
   KNRL_K_NTH_ADJ : ALIAS FOR O[19].0;
   KNRL_K_STH_ADJ : ALIAS FOR O[19].1;
   KNRL_N_AUTO : ALIAS FOR N14[250].0;
   KNRL_N_MANL : ALIAS FOR N14[251].0;
   KNRL_S_AUTO : ALIAS FOR N14[250].1;
   KNRL_S_MANL : ALIAS FOR N14[251].1;
   KNRL_T_NTH_ADJ : ALIAS FOR O[22].0;
   KNRL_T_STH_ADJ : ALIAS FOR O[22].1;
   LEHR_SPEED : ALIAS FOR N20[1];
   LINE_SPEED : ALIAS FOR N20[3];
   M2_ALM_HORN_RLY : ALIAS FOR O[9].3;
   M2_ALM_RESET : ALIAS FOR I[2].9;
   M2_ALM_SILENCE : ALIAS FOR I[2].8;
   M2_AMBER_STKLTE : ALIAS FOR O[9].6;
   M2_BLUE_STKLTE : ALIAS FOR O[9].5;
   M2_CM07N_HZIMP : DINT := 1853;   // This compute statement was created to allow speed control on M2 CM07N; 28Mar2019,AAC.
   M2_CM07N_Lehr_Speed : DINT := 71;   // This compute statement was created to allow speed control for Lehr Speed on M2 CM07N; 28Mar2019,AAC.
   M2_CM07N_Slip_Comp : DINT := 1160;
   M2_CM07N_Trim_Speed : DINT := 243;   // This compute statement was created to allow Trim speed control on M2 CM07N; 28Mar2019,AAC.
   M2_DC_INPWR : ALIAS FOR I[2].2;
   M2_DC_OUTPWR : ALIAS FOR I[2].3;
   M2_DC_PS1 : ALIAS FOR I[2].6;
   M2_DC_PS2 : ALIAS FOR I[2].7;
   M2_DRV_CONT_ON : ALIAS FOR I[2].1;
   M2_DRV_FLT_LMP : ALIAS FOR O[9].0;
   M2_ESTOP : ALIAS FOR I[2].10;
   M2_ESTOPPWR : ALIAS FOR I[2].5;
   M2_FLT_RES_RLY : ALIAS FOR O[9].1;
   M2_RED_STKLTE : ALIAS FOR O[9].4;
   M301_M1_TD_DR : AXIS_CIP_DRIVE; {access Read Only}
   M301_M1_TK_DR : AXIS_CIP_DRIVE; {access Read Only}
   M301_M2_TD_DR : AXIS_CIP_DRIVE; {access Read Only}
   M301_M2_TK_DR : AXIS_CIP_DRIVE; {access Read Only}
   M302_M1_TD_DR : AXIS_CIP_DRIVE; {access Read Only}
   M302_M1_TK_DR : AXIS_CIP_DRIVE; {access Read Only}
   M302_M2_TD_DR : AXIS_CIP_DRIVE; {access Read Only}
   M302_M2_TK_DR : AXIS_CIP_DRIVE; {access Read Only}
   M302SpeedUp : MAC_SpeedUp := (OSR_xAccDecHighForThicknessLow := 1, INPUT_xControlSnap1 := 1, INPUT_xControlSnap2 := 1, INPUT_rRealSpeedInAcc_mm_min := 11167.0, INPUT_dDecRamp_m_s2 := 1.2, AUX_dMaxMissSnap := 2, AUX_dMaxCapLength_cmm := 700000, AUX_dControlSnapLimit_cmm := 30000, AUX_dConveyorLength_cmm := 712500, AUX_dLastDataReceived := 905816, AUX_dDimensionCapCreation_cmm := 49104, AUX_dDimensionCapMissSnap_cmm := 49104, AUX_dLastIndexTailSnap := 6, AUX_dFirstIndexHeadSnap := 6, AUX_dLastConvoyTailPos_cmm := 162595, AUX_dConvoyGlassLength_cmm := 270000, AUX_dMaxConvoyLength_cmm := 360000, AUX_dSymmetricGap_cmm := 15000, AUX_dConvoyLengthTarget_cmm := 300000, AUX_dNumCapsInConvoy := 3, AUX_dManualSideLegWidth_cmm := 344000, AUX_dStandardGap_cmm := 15000, rgxReqAcc := 28, AUX_rLehrStepInc_cmm := 372.23334, tmON_TimeControlSnap[0].PRE := 30000, tmON_TimeControlSnap[1].PRE := 30000, tmON_GapCount.PRE := 339, tSearchPlate.rgdHeadPointer[0] := 6, tSearchPlate.rgdTailPointer[0] := 6, tSearchPlate.rgdHead_cmm[0] := 422595, tSearchPlate.rgdTail_cmm[0] := 162595, tSearchPlate.rgxHead := 1, tSearchPlate.rgxTail := 1, tSearchPlate.xHeadPresence := 1, tSearchPlate.xTailPresence := 1); {access None}
   M302SpeedUp_ALM : MAC_SpeedUp_ALM; {access Read Only}
        .rgxFault.1   // M302.Plate length error
        .rgxFault.0   // M302.Missing snap error
        .rgxFault.2   // M302.Plate length over specifications
        .rgxWarning.0   // M302.Timeout Break-out control photocell #1
        .rgxWarning.1   // M302.Timeout Break-out control photocell #2
   M302SpeedUp_HMR : MAC_SpeedUp_HMR := (xControlSnap1 := 1, xControlSnap2 := 1, dControlSnapEnabled := 1, rgdStateSensor[0] := 1, rgdStateSensor[1] := 1); {access Read Only}
   M302SpeedUp_HMW : MAC_SpeedUp_HMW;
   M302SpeedUp_tmON_ProtSnap : TIMER := (PRE := 50); {access Read Only}
   M302SpeedUp_xFirstScanProtSnap : BOOL; {access Read Only}
   M303_dHalfWidthDifference : DINT := 2900; {access Read Only}
   M303_M1_TD_DR : AXIS_CIP_DRIVE; {access Read Only}
   M303_M1_TK_DR : AXIS_CIP_DRIVE; {access Read Only}
   M303_M2_TD_DR : AXIS_CIP_DRIVE; {access Read Only}
   M303_M2_TK_DR : AXIS_CIP_DRIVE; {access Read Only}
   M304_M1_TD_DR : AXIS_CIP_DRIVE; {access Read Only}
   M304_M1_TK_DR : AXIS_CIP_DRIVE; {access Read Only}
   M304_M2_TD_DR : AXIS_CIP_DRIVE; {access Read Only}
   M304_M2_TK_DR : AXIS_CIP_DRIVE; {access Read Only}
   M305_M1_TD_DR : AXIS_CIP_DRIVE; {access Read Only}
   M305_M1_TK_DR : AXIS_CIP_DRIVE; {access Read Only}
   M305_M2_TD_DR : AXIS_CIP_DRIVE; {access Read Only}
   M305_M2_TK_DR : AXIS_CIP_DRIVE; {access Read Only}
   M306_M1_TD_DR : AXIS_CIP_DRIVE; {access Read Only}
   M306_M1_TK_DR : AXIS_CIP_DRIVE; {access Read Only}
   M306_M2_TD_DR : AXIS_CIP_DRIVE; {access Read Only}
   M306_M2_TK_DR : AXIS_CIP_DRIVE; {access Read Only}
   M307A_M1_DR : AXIS_CIP_DRIVE; {access Read Only}
   M307A_M2_DR : AXIS_CIP_DRIVE; {access Read Only}
   M307A_M3_DR : AXIS_CIP_DRIVE; {access Read Only}
   M307A_M4_DR : AXIS_CIP_DRIVE; {access Read Only}
   M307ASpeedUp : MAC_SpeedUp := (ST_xConditionOKChangeSpeed := 1, ST_xPlateComing := 1, OSR_xNewData := 1, AUX_dConveyorLength_cmm := 800000, AUX_dDimensionCapCreation_cmm := 44064, AUX_dLastConvoyTailPos_cmm := 3428619, rgxReqAcc := 4, AUX_rLehrStepInc_cmm := 1295.6, tmON_TimeControlSnap[0].PRE := 30000, tmON_TimeControlSnap[1].PRE := 30000, tSearchPlate.rgdHeadPointer[0] := 7, tSearchPlate.rgdHead_cmm[0] := 2669958, tSearchPlate.rgxHead := 1, tSearchPlate.xHeadPresence := 1); {access None}
   M307ASpeedUp_ALM : MAC_SpeedUp_ALM; {access Read Only}
   M307ASpeedUp_HMR : MAC_SpeedUp_HMR := (xControlSnap1 := 1, xControlSnap2 := 1, rgdStateSensor[0] := 1, rgdStateSensor[1] := 1); {access Read Only}
   M307ASpeedUp_HMW : MAC_SpeedUp_HMW;
   M307B_M1_DR : AXIS_CIP_DRIVE; {access Read Only}
   M307C_M1_DR : AXIS_CIP_DRIVE; {access Read Only}
   M307D_M1_DR : AXIS_CIP_DRIVE; {access Read Only}
   M307E_M1_DR : AXIS_CIP_DRIVE; {access Read Only}
   M307F_M1_DR : AXIS_CIP_DRIVE; {access Read Only}
   M30xTrimDeck : MAC_TrimmingDeck[5]; {access None}
        [0]   // M302
        [1]   // M303
        [2]   // M304
        [3]   // M305
        [4]   // M306
   M30xTrimDeck_ALM : MAC_TrimmingDeck_ALM[5]; {access Read Only}
        [1]   // M303
        [2]   // M304
        [0]   // M302
        [0].rgxStoppingFault_M[0].x1   // M302.Drive error trim deck operator side
        [3]   // M305
        [4]   // M306
        [0].rgxStoppingFault_M[0].x0   // M302.Protection motor trim deck operator side
        [0].rgxStoppingFault_M[0].x2   // M302.Drive feedback error trim deck operator side
        [0].rgxStoppingFault_M[0].x3   // M302.Local safety switch trim deck operator side
        [0].rgxStoppingFault_M[0].x4   // M302.Motor thermal probe trim deck operator side
        [0].rgxStoppingFault_M[0].x5   // M302.Braking resistor fault trim deck operator side
        [0].rgxStoppingFault_M[0].x6   // M302.Encoder error trim deck operator side
        [0].rgxStoppingFault_M[1].x0   // M302.Protection motor trim deck opposite operator side
        [0].rgxStoppingFault_M[1].x1   // M302.Drive error trim deck opposite operator side
        [0].rgxStoppingFault_M[1].x2   // M302.Drive feedback error trim deck opposite operator side
        [0].rgxStoppingFault_M[1].x3   // M302.Local safety switch trim deck opposite operator side
        [0].rgxStoppingFault_M[1].x4   // M302.Motor thermal probe trim deck opposite operator side
        [0].rgxStoppingFault_M[1].x5   // M302.Braking resistor fault trim deck opposite operator side
        [0].rgxStoppingFault_M[1].x6   // M302.Encoder error trim deck opposite operator side
        [1].rgxStoppingFault_M[0].x0   // M303.Protection motor trim deck operator side
        [1].rgxStoppingFault_M[1].x0   // M303.Protection motor trim deck opposite operator side
        [1].rgxStoppingFault_M[0].x1   // M303.Drive error trim deck operator side
        [3].rgxStoppingFault_M[0].x1   // M305.Drive error trim deck operator side
        [2].rgxStoppingFault_M[0].x1   // M304.Drive error trim deck operator side
        [2].rgxStoppingFault_M[1].x1   // M304.Drive error trim deck opposite operator side
        [2].rgxStoppingFault_M[0].x0   // M304.Protection motor trim deck operator side
        [2].rgxStoppingFault_M[1].x0   // M304.Protection motor trim deck opposite operator side
        [1].rgxStoppingFault_M[0].x3   // M303.Local safety switch trim deck operator side
        [1].rgxStoppingFault_M[0].x2   // M303.Drive feedback error trim deck operator side
        [1].rgxStoppingFault_M[1].x3   // M303.Local safety switch trim deck opposite operator side
        [1].rgxStoppingFault_M[1].x1   // M303.Drive error trim deck opposite operator side
        [1].rgxStoppingFault_M[1].x2   // M303.Drive feedback error trim deck opposite operator side
        [1].rgxStoppingFault_M[1].x4   // M303.Motor thermal probe trim deck opposite operator side
        [1].rgxStoppingFault_M[1].x5   // M303.Braking resistor fault trim deck opposite operator side
        [1].rgxStoppingFault_M[1].x6   // M303.Encoder error trim deck opposite operator side
        [1].rgxStoppingFault_M[0].x4   // M303.Motor thermal probe trim deck operator side
        [1].rgxStoppingFault_M[0].x5   // M303.Braking resistor fault trim deck operator side
        [1].rgxStoppingFault_M[0].x6   // M303.Encoder error trim deck operator side
        [2].rgxStoppingFault_M[0].x4   // M304.Motor thermal probe trim deck operator side
        [2].rgxStoppingFault_M[1].x4   // M304.Motor thermal probe trim deck opposite operator side
        [2].rgxStoppingFault_M[1].x2   // M304.Drive feedback error trim deck opposite operator side
        [2].rgxStoppingFault_M[1].x3   // M304.Local safety switch trim deck opposite operator side
        [2].rgxStoppingFault_M[1].x5   // M304.Braking resistor fault trim deck opposite operator side
        [2].rgxStoppingFault_M[1].x6   // M304.Encoder error trim deck opposite operator side
        [2].rgxStoppingFault_M[0].x6   // M304.Encoder error trim deck operator side
        [2].rgxStoppingFault_M[0].x2   // M304.Drive feedback error trim deck operator side
        [2].rgxStoppingFault_M[0].x3   // M304.Local safety switch trim deck operator side
        [2].rgxStoppingFault_M[0].x5   // M304.Braking resistor fault trim deck operator side
        [3].rgxStoppingFault_M[0].x0   // M305.Protection motor trim deck operator side
        [3].rgxStoppingFault_M[1].x0   // M305.Protection motor trim deck opposite operator side
        [3].rgxStoppingFault_M[1].x1   // M305.Drive error trim deck opposite operator side
        [3].rgxStoppingFault_M[1].x2   // M305.Drive feedback error trim deck opposite operator side
        [3].rgxStoppingFault_M[1].x3   // M305.Local safety switchtrim deck opposite operator side
        [3].rgxStoppingFault_M[1].x4   // M305.Motor thermal probe trim deck opposite operator side
        [3].rgxStoppingFault_M[1].x5   // M305.Braking resistor fault trim deck opposite operator side
        [3].rgxStoppingFault_M[1].x6   // M305.Encoder error trim deck opposite operator side
        [3].rgxStoppingFault_M[0].x2   // M305.Drive feddback error trim deck operator side
        [3].rgxStoppingFault_M[0].x3   // M305.Local safety switch trim deck operator side
        [3].rgxStoppingFault_M[0].x4   // M305.Motor thermal probe trim deck operator side
        [3].rgxStoppingFault_M[0].x5   // M305.Braking resistor fault trim deck operator side
        [3].rgxStoppingFault_M[0].x6   // M305.Encoder error trim deck operator side
        [4].rgxStoppingFault_M[0].x0   // M306.Protection motor trim deck operator side
        [4].rgxStoppingFault_M[0].x1   // M306.Drive error trim deck operator side
        [4].rgxStoppingFault_M[0].x2   // M306.Drive feedback error trim deck operator side
        [4].rgxStoppingFault_M[1].x1   // M306.Drive error trim deck opposite operator side
        [4].rgxStoppingFault_M[1].x2   // M306.Drive feedback error trim deck opposite operator side
        [4].rgxStoppingFault_M[1].x0   // M306.Protection motor trim deck opposite operator side
        [4].rgxStoppingFault_M[1].x3   // M306.Local safety switch trim deck opposite operator side
        [4].rgxStoppingFault_M[1].x4   // M306.Motor thermal probe trim deck opposite operator side
        [4].rgxStoppingFault_M[1].x5   // M306.Braking resistor fault trim deck opposite operator side
        [4].rgxStoppingFault_M[1].x6   // M306.Encoder error trim deck opposite operator side
        [4].rgxStoppingFault_M[0].x3   // M306.Local safety switch trim deck operator side
        [4].rgxStoppingFault_M[0].x4   // M306.Motor thermal probe trim deck operator side
        [4].rgxStoppingFault_M[0].x5   // M306.Braking resistor fault trim deck operator side
        [4].rgxStoppingFault_M[0].x6   // M306.Encoder error trim deck operator side
   M30xTrimDeck_DATA : UDT_ConvoyCap_ZC[5];
        [4]   // Cap data M306
        [0]   // Cap data M302
        [1]   // Cap data M303
        [2]   // Cap data M304
        [3]   // Cap data M305
   M30xTrimDeck_HMR : MAC_TrimmingDeck_HMR[5] := ([0].xControlWidthEnabled := 1, [0].xControlWanderEnabled := 1, [0].xCulletEdgeEnabled := 1, [0].xOpeningOnCleaningEnabled := 1, [0].rgdState[0] := 1, [0].rgdState[1] := 1, [0].dGrossWidthInProgress_cmm := 377400, [0].dNetWidthInProgress_cmm := 360000, [0].dCutWanderInProgress_cmm := -3930, [0].rgdTarget_cmm[0] := 185430, [0].rgdTarget_cmm[1] := 181570, [0].rgdPosition_cmm[0] := 185399, [0].rgdPosition_cmm[1] := 181500, [0].rgdOffsetEachSide_cmm[0] := 1500, [0].rgdOffsetEachSide_cmm[1] := 5500, [0].dDistBetweenSides_cmm := 366899); {access Read Only}
        [0]   // M302
        [1]   // M303
        [2]   // M304
        [3]   // M305
        [4]   // M306
   M30xTrimDeck_HMW : MAC_TrimmingDeck_HMW[5] := ([0].xEnableDisableCulletEdge := 1, [0].dOffsetOpSide_cmm := 1500, [0].dOffsetOppOpSide_cmm := 5500);
        [0]   // M302
        [1]   // M303
        [2]   // M304
        [3]   // M305
        [4]   // M306
   M30xTrimDeck_IN_MOTION : MAC_TrimmingDeck_IN_MOTION[5] := ([0].DR_MAJ_M[0].FLAGS := 33554432, [0].DR_MAJ_M[1].FLAGS := 33554432, [0].DR_MAM_M[0].FLAGS := 704643072, [0].DR_MAM_M[0].DN := 1, [0].DR_MAM_M[0].PC := 1, [0].DR_MAM_M[1].FLAGS := 704643072, [0].DR_MAM_M[1].DN := 1, [0].DR_MAM_M[1].PC := 1, [0].DR_MAS_M[0].FLAGS := -1442840576, [0].DR_MAS_M[0].EN := 1, [0].DR_MAS_M[0].DN := 1, [0].DR_MAS_M[0].PC := 1, [0].DR_MAS_M[1].FLAGS := -1442840576, [0].DR_MAS_M[1].EN := 1, [0].DR_MAS_M[1].DN := 1, [0].DR_MAS_M[1].PC := 1); {access None}
   M30xTrimDeck_OUT_MOTION : MAC_TrimmingDeck_OUT_MOTION[5] := ([0].DR_MSO_M[0].FLAGS := -1610612736, [0].DR_MSO_M[0].EN := 1, [0].DR_MSO_M[0].DN := 1, [0].DR_MSO_M[0].STATE := 1, [0].DR_MSO_M[1].FLAGS := -1610612736, [0].DR_MSO_M[1].EN := 1, [0].DR_MSO_M[1].DN := 1, [0].DR_MSO_M[1].STATE := 1, [0].DR_MSF_M[0].FLAGS := 570425344, [0].DR_MSF_M[0].DN := 1, [0].DR_MSF_M[0].STATUS := 2, [0].DR_MSF_M[0].STATE := 1, [0].DR_MSF_M[1].FLAGS := 570425344, [0].DR_MSF_M[1].DN := 1, [0].DR_MSF_M[1].STATUS := 2, [0].DR_MSF_M[1].STATE := 1, [0].DR_MASR_M[0].FLAGS := 536870912, [0].DR_MASR_M[0].DN := 1, [0].DR_MASR_M[0].STATE := 1, [0].DR_MASR_M[1].FLAGS := 536870912, [0].DR_MASR_M[1].DN := 1, [0].DR_MASR_M[1].STATE := 1, [0].DR_MAJ_M[0].FLAGS := 33554432, [0].DR_MAJ_M[1].FLAGS := 33554432, [0].DR_MAM_M[0].FLAGS := 704643072, [0].DR_MAM_M[0].DN := 1, [0].DR_MAM_M[0].PC := 1, [0].DR_MAM_M[1].FLAGS := 704643072, [0].DR_MAM_M[1].DN := 1, [0].DR_MAM_M[1].PC := 1, [0].DR_MCD_M[0].FLAGS := 33554432, [0].DR_MCD_M[1].FLAGS := 33554432, [0].DR_MAS_M[0].FLAGS := -1442840576, [0].DR_MAS_M[0].EN := 1, [0].DR_MAS_M[0].DN := 1, [0].DR_MAS_M[0].PC := 1, [0].DR_MAS_M[1].FLAGS := -1442840576, [0].DR_MAS_M[1].EN := 1, [0].DR_MAS_M[1].DN := 1, [0].DR_MAS_M[1].PC := 1, [0].DR_MAH_M[0].FLAGS := 33554432, [0].DR_MAH_M[1].FLAGS := 33554432); {access None}